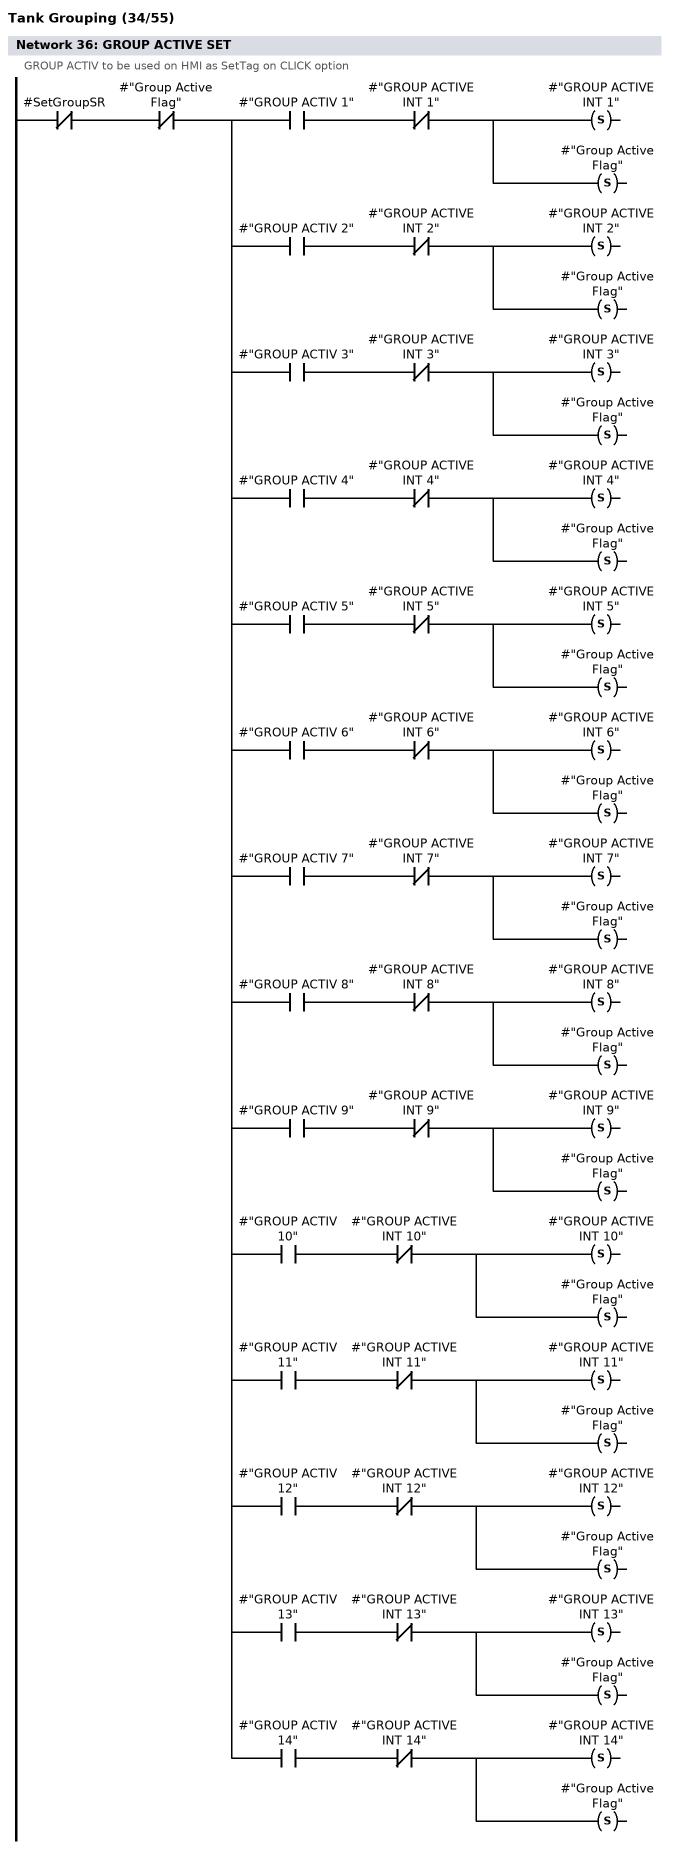
   RUNG wire#powerrail
      I_Contact( #SetGroupSR )
      I_Contact( #"Group Active Flag" )
      wire#w1
      Contact( #"GROUP ACTIV 1" )
      I_Contact( #"GROUP ACTIVE INT 1" )
      wire#w2
      S_Coil( #"GROUP ACTIVE INT 1" )
   END_RUNG
   RUNG wire#w2
      S_Coil( #"Group Active Flag" )
   END_RUNG
   RUNG wire#w1
      Contact( #"GROUP ACTIV 2" )
      I_Contact( #"GROUP ACTIVE INT 2" )
      wire#w3
      S_Coil( #"GROUP ACTIVE INT 2" )
   END_RUNG
   RUNG wire#w3
      S_Coil( #"Group Active Flag" )
   END_RUNG
   RUNG wire#w1
      Contact( #"GROUP ACTIV 3" )
      I_Contact( #"GROUP ACTIVE INT 3" )
      wire#w4
      S_Coil( #"GROUP ACTIVE INT 3" )
   END_RUNG
   RUNG wire#w4
      S_Coil( #"Group Active Flag" )
   END_RUNG
   RUNG wire#w1
      Contact( #"GROUP ACTIV 4" )
      I_Contact( #"GROUP ACTIVE INT 4" )
      wire#w5
      S_Coil( #"GROUP ACTIVE INT 4" )
   END_RUNG
   RUNG wire#w5
      S_Coil( #"Group Active Flag" )
   END_RUNG
   RUNG wire#w1
      Contact( #"GROUP ACTIV 5" )
      I_Contact( #"GROUP ACTIVE INT 5" )
      wire#w6
      S_Coil( #"GROUP ACTIVE INT 5" )
   END_RUNG
   RUNG wire#w6
      S_Coil( #"Group Active Flag" )
   END_RUNG
   RUNG wire#w1
      Contact( #"GROUP ACTIV 6" )
      I_Contact( #"GROUP ACTIVE INT 6" )
      wire#w7
      S_Coil( #"GROUP ACTIVE INT 6" )
   END_RUNG
   RUNG wire#w7
      S_Coil( #"Group Active Flag" )
   END_RUNG
   RUNG wire#w1
      Contact( #"GROUP ACTIV 7" )
      I_Contact( #"GROUP ACTIVE INT 7" )
      wire#w8
      S_Coil( #"GROUP ACTIVE INT 7" )
   END_RUNG
   RUNG wire#w8
      S_Coil( #"Group Active Flag" )
   END_RUNG
   RUNG wire#w1
      Contact( #"GROUP ACTIV 8" )
      I_Contact( #"GROUP ACTIVE INT 8" )
      wire#w9
      S_Coil( #"GROUP ACTIVE INT 8" )
   END_RUNG
   RUNG wire#w9
      S_Coil( #"Group Active Flag" )
   END_RUNG
   RUNG wire#w1
      Contact( #"GROUP ACTIV 9" )
      I_Contact( #"GROUP ACTIVE INT 9" )
      wire#w10
      S_Coil( #"GROUP ACTIVE INT 9" )
   END_RUNG
   RUNG wire#w10
      S_Coil( #"Group Active Flag" )
   END_RUNG
   RUNG wire#w1
      Contact( #"GROUP ACTIV 10" )
      I_Contact( #"GROUP ACTIVE INT 10" )
      wire#w11
      S_Coil( #"GROUP ACTIVE INT 10" )
   END_RUNG
   RUNG wire#w11
      S_Coil( #"Group Active Flag" )
   END_RUNG
   RUNG wire#w1
      Contact( #"GROUP ACTIV 11" )
      I_Contact( #"GROUP ACTIVE INT 11" )
      wire#w12
      S_Coil( #"GROUP ACTIVE INT 11" )
   END_RUNG
   RUNG wire#w12
      S_Coil( #"Group Active Flag" )
   END_RUNG
   RUNG wire#w1
      Contact( #"GROUP ACTIV 12" )
      I_Contact( #"GROUP ACTIVE INT 12" )
      wire#w13
      S_Coil( #"GROUP ACTIVE INT 12" )
   END_RUNG
   RUNG wire#w13
      S_Coil( #"Group Active Flag" )
   END_RUNG
   RUNG wire#w1
      Contact( #"GROUP ACTIV 13" )
      I_Contact( #"GROUP ACTIVE INT 13" )
      wire#w14
      S_Coil( #"GROUP ACTIVE INT 13" )
   END_RUNG
   RUNG wire#w14
      S_Coil( #"Group Active Flag" )
   END_RUNG
   RUNG wire#w1
      Contact( #"GROUP ACTIV 14" )
      I_Contact( #"GROUP ACTIVE INT 14" )
      wire#w15
      S_Coil( #"GROUP ACTIVE INT 14" )
   END_RUNG
   RUNG wire#w15
      S_Coil( #"Group Active Flag" )
   END_RUNG
   // the same network as SCL:
   #_w1 := NOT #SetGroupSR AND NOT #"Group Active Flag";
   #_w2 := #_w1 AND #"GROUP ACTIV 1" AND NOT #"GROUP ACTIVE INT 1";
   IF #_w2 THEN
       #"GROUP ACTIVE INT 1" := TRUE;
       #"Group Active Flag" := TRUE;
   END_IF;
   #_w3 := #_w1 AND #"GROUP ACTIV 2" AND NOT #"GROUP ACTIVE INT 2";
   IF #_w3 THEN
       #"GROUP ACTIVE INT 2" := TRUE;
       #"Group Active Flag" := TRUE;
   END_IF;
   #_w4 := #_w1 AND #"GROUP ACTIV 3" AND NOT #"GROUP ACTIVE INT 3";
   IF #_w4 THEN
       #"GROUP ACTIVE INT 3" := TRUE;
       #"Group Active Flag" := TRUE;
   END_IF;
   #_w5 := #_w1 AND #"GROUP ACTIV 4" AND NOT #"GROUP ACTIVE INT 4";
   IF #_w5 THEN
       #"GROUP ACTIVE INT 4" := TRUE;
       #"Group Active Flag" := TRUE;
   END_IF;
   #_w6 := #_w1 AND #"GROUP ACTIV 5" AND NOT #"GROUP ACTIVE INT 5";
   IF #_w6 THEN
       #"GROUP ACTIVE INT 5" := TRUE;
       #"Group Active Flag" := TRUE;
   END_IF;
   #_w7 := #_w1 AND #"GROUP ACTIV 6" AND NOT #"GROUP ACTIVE INT 6";
   IF #_w7 THEN
       #"GROUP ACTIVE INT 6" := TRUE;
       #"Group Active Flag" := TRUE;
   END_IF;
   #_w8 := #_w1 AND #"GROUP ACTIV 7" AND NOT #"GROUP ACTIVE INT 7";
   IF #_w8 THEN
       #"GROUP ACTIVE INT 7" := TRUE;
       #"Group Active Flag" := TRUE;
   END_IF;
   #_w9 := #_w1 AND #"GROUP ACTIV 8" AND NOT #"GROUP ACTIVE INT 8";
   IF #_w9 THEN
       #"GROUP ACTIVE INT 8" := TRUE;
       #"Group Active Flag" := TRUE;
   END_IF;
   #_w10 := #_w1 AND #"GROUP ACTIV 9" AND NOT #"GROUP ACTIVE INT 9";
   IF #_w10 THEN
       #"GROUP ACTIVE INT 9" := TRUE;
       #"Group Active Flag" := TRUE;
   END_IF;
   #_w11 := #_w1 AND #"GROUP ACTIV 10" AND NOT #"GROUP ACTIVE INT 10";
   IF #_w11 THEN
       #"GROUP ACTIVE INT 10" := TRUE;
       #"Group Active Flag" := TRUE;
   END_IF;
   #_w12 := #_w1 AND #"GROUP ACTIV 11" AND NOT #"GROUP ACTIVE INT 11";
   IF #_w12 THEN
       #"GROUP ACTIVE INT 11" := TRUE;
       #"Group Active Flag" := TRUE;
   END_IF;
   #_w13 := #_w1 AND #"GROUP ACTIV 12" AND NOT #"GROUP ACTIVE INT 12";
   IF #_w13 THEN
       #"GROUP ACTIVE INT 12" := TRUE;
       #"Group Active Flag" := TRUE;
   END_IF;
   #_w14 := #_w1 AND #"GROUP ACTIV 13" AND NOT #"GROUP ACTIVE INT 13";
   IF #_w14 THEN
       #"GROUP ACTIVE INT 13" := TRUE;
       #"Group Active Flag" := TRUE;
   END_IF;
   #_w15 := #_w1 AND #"GROUP ACTIV 14" AND NOT #"GROUP ACTIVE INT 14";
   IF #_w15 THEN
       #"GROUP ACTIVE INT 14" := TRUE;
       #"Group Active Flag" := TRUE;
   END_IF;
END_REGION

REGION Network 37: Group Active Flag Reset
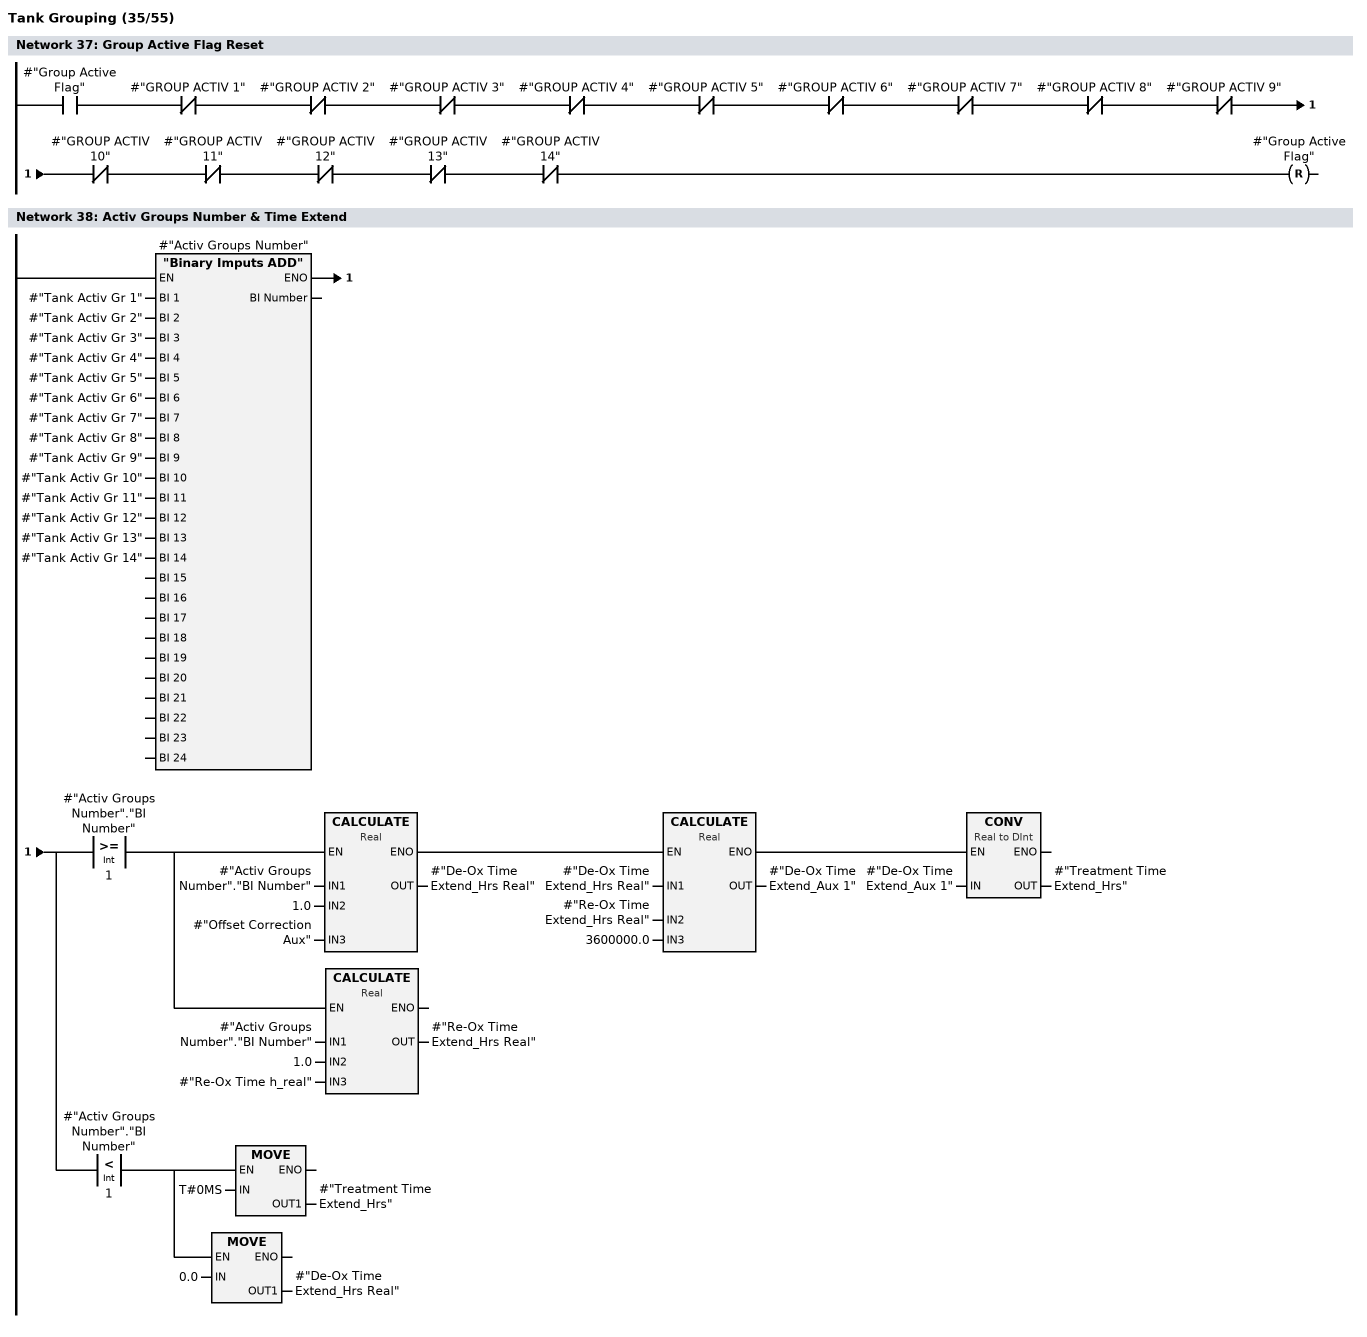
   RUNG wire#powerrail
      Contact( #"Group Active Flag" )
      I_Contact( #"GROUP ACTIV 1" )
      I_Contact( #"GROUP ACTIV 2" )
      I_Contact( #"GROUP ACTIV 3" )
      I_Contact( #"GROUP ACTIV 4" )
      I_Contact( #"GROUP ACTIV 5" )
      I_Contact( #"GROUP ACTIV 6" )
      I_Contact( #"GROUP ACTIV 7" )
      I_Contact( #"GROUP ACTIV 8" )
      I_Contact( #"GROUP ACTIV 9" )
      I_Contact( #"GROUP ACTIV 10" )
      I_Contact( #"GROUP ACTIV 11" )
      I_Contact( #"GROUP ACTIV 12" )
      I_Contact( #"GROUP ACTIV 13" )
      I_Contact( #"GROUP ACTIV 14" )
      R_Coil( #"Group Active Flag" )
   END_RUNG
   // the same network as SCL:
   IF #"Group Active Flag" AND NOT #"GROUP ACTIV 1" AND NOT #"GROUP ACTIV 2" AND NOT #"GROUP ACTIV 3" AND NOT #"GROUP ACTIV 4" AND NOT #"GROUP ACTIV 5" AND NOT #"GROUP ACTIV 6" AND NOT #"GROUP ACTIV 7" AND NOT #"GROUP ACTIV 8" AND NOT #"GROUP ACTIV 9" AND NOT #"GROUP ACTIV 10" AND NOT #"GROUP ACTIV 11" AND NOT #"GROUP ACTIV 12" AND NOT #"GROUP ACTIV 13" AND NOT #"GROUP ACTIV 14" THEN
       #"Group Active Flag" := FALSE;
   END_IF;
END_REGION

REGION Network 38: Activ Groups Number & Time Extend
   RUNG wire#powerrail
      #"Activ Groups Number"("BI 1" := #"Tank Activ Gr 1", "BI 2" := #"Tank Activ Gr 2", "BI 3" := #"Tank Activ Gr 3", "BI 4" := #"Tank Activ Gr 4", "BI 5" := #"Tank Activ Gr 5", "BI 6" := #"Tank Activ Gr 6", "BI 7" := #"Tank Activ Gr 7", "BI 8" := #"Tank Activ Gr 8", "BI 9" := #"Tank Activ Gr 9", "BI 10" := #"Tank Activ Gr 10", "BI 11" := #"Tank Activ Gr 11", "BI 12" := #"Tank Activ Gr 12", "BI 13" := #"Tank Activ Gr 13", "BI 14" := #"Tank Activ Gr 14", "BI 15" :=, "BI 16" :=, "BI 17" :=, "BI 18" :=, "BI 19" :=, "BI 20" :=, "BI 21" :=, "BI 22" :=, "BI 23" :=, "BI 24" :=, "BI Number" =>)
      wire#w1
      { S7_Templates := "SrcType := Int" } GE_Contact(in1 := #"Activ Groups Number"."BI Number", in2 := 1)
      wire#w2
      { S7_Templates := "SrcType := Real"; S7_Expression := "IN3*(IN1-IN2)" } Calculate(in1 := #"Activ Groups Number"."BI Number", in2 := 1.0, in3 := #"Offset Correction Aux", out => #"De-Ox Time Extend_Hrs Real")
      { S7_Templates := "SrcType := Real"; S7_Expression := "(IN1+IN2)*IN3" } Calculate(in1 := #"De-Ox Time Extend_Hrs Real", in2 := #"Re-Ox Time Extend_Hrs Real", in3 := 3600000.0, out => #"De-Ox Time Extend_Aux 1")
      { S7_Templates := "[SrcType := Real, DestType := DInt]" } Convert(in := #"De-Ox Time Extend_Aux 1", out => #"Treatment Time Extend_Hrs")
   END_RUNG
   RUNG wire#w2
      { S7_Templates := "SrcType := Real"; S7_Expression := "IN3*(IN1-IN2)" } Calculate(in1 := #"Activ Groups Number"."BI Number", in2 := 1.0, in3 := #"Re-Ox Time h_real", out => #"Re-Ox Time Extend_Hrs Real")
   END_RUNG
   RUNG wire#w1
      { S7_Templates := "SrcType := Int" } LT_Contact(in1 := #"Activ Groups Number"."BI Number", in2 := 1)
      wire#w3
      Move(in := T#0MS, out1 => #"Treatment Time Extend_Hrs")
   END_RUNG
   RUNG wire#w3
      Move(in := 0.0, out1 => #"De-Ox Time Extend_Hrs Real")
   END_RUNG
   // the same network as SCL:
   #"Activ Groups Number"("BI 1" := #"Tank Activ Gr 1",   // "Binary Imputs ADD"
                          "BI 2" := #"Tank Activ Gr 2",
                          "BI 3" := #"Tank Activ Gr 3",
                          "BI 4" := #"Tank Activ Gr 4",
                          "BI 5" := #"Tank Activ Gr 5",
                          "BI 6" := #"Tank Activ Gr 6",
                          "BI 7" := #"Tank Activ Gr 7",
                          "BI 8" := #"Tank Activ Gr 8",
                          "BI 9" := #"Tank Activ Gr 9",
                          "BI 10" := #"Tank Activ Gr 10",
                          "BI 11" := #"Tank Activ Gr 11",
                          "BI 12" := #"Tank Activ Gr 12",
                          "BI 13" := #"Tank Activ Gr 13",
                          "BI 14" := #"Tank Activ Gr 14",
                          ENO => #_w1);
   IF #_w1 AND (#"Activ Groups Number"."BI Number" >= 1) THEN
       #"De-Ox Time Extend_Hrs Real" := #"Offset Correction Aux"*(#"Activ Groups Number"."BI Number"-1.0);
       #"De-Ox Time Extend_Aux 1" := (#"De-Ox Time Extend_Hrs Real"+#"Re-Ox Time Extend_Hrs Real")*3600000.0;
       #"Treatment Time Extend_Hrs" := REAL_TO_DINT(#"De-Ox Time Extend_Aux 1");
       #"Re-Ox Time Extend_Hrs Real" := #"Re-Ox Time h_real"*(#"Activ Groups Number"."BI Number"-1.0);
   END_IF;
   IF #_w1 AND (#"Activ Groups Number"."BI Number" < 1) THEN
       #"Treatment Time Extend_Hrs" := T#0MS;
       #"De-Ox Time Extend_Hrs Real" := 0.0;
   END_IF;
END_REGION

REGION Network 39: GROUP ACTIVE RESET
   // GROUP ACTIV to be used on HMI as SetTag on CLICK option
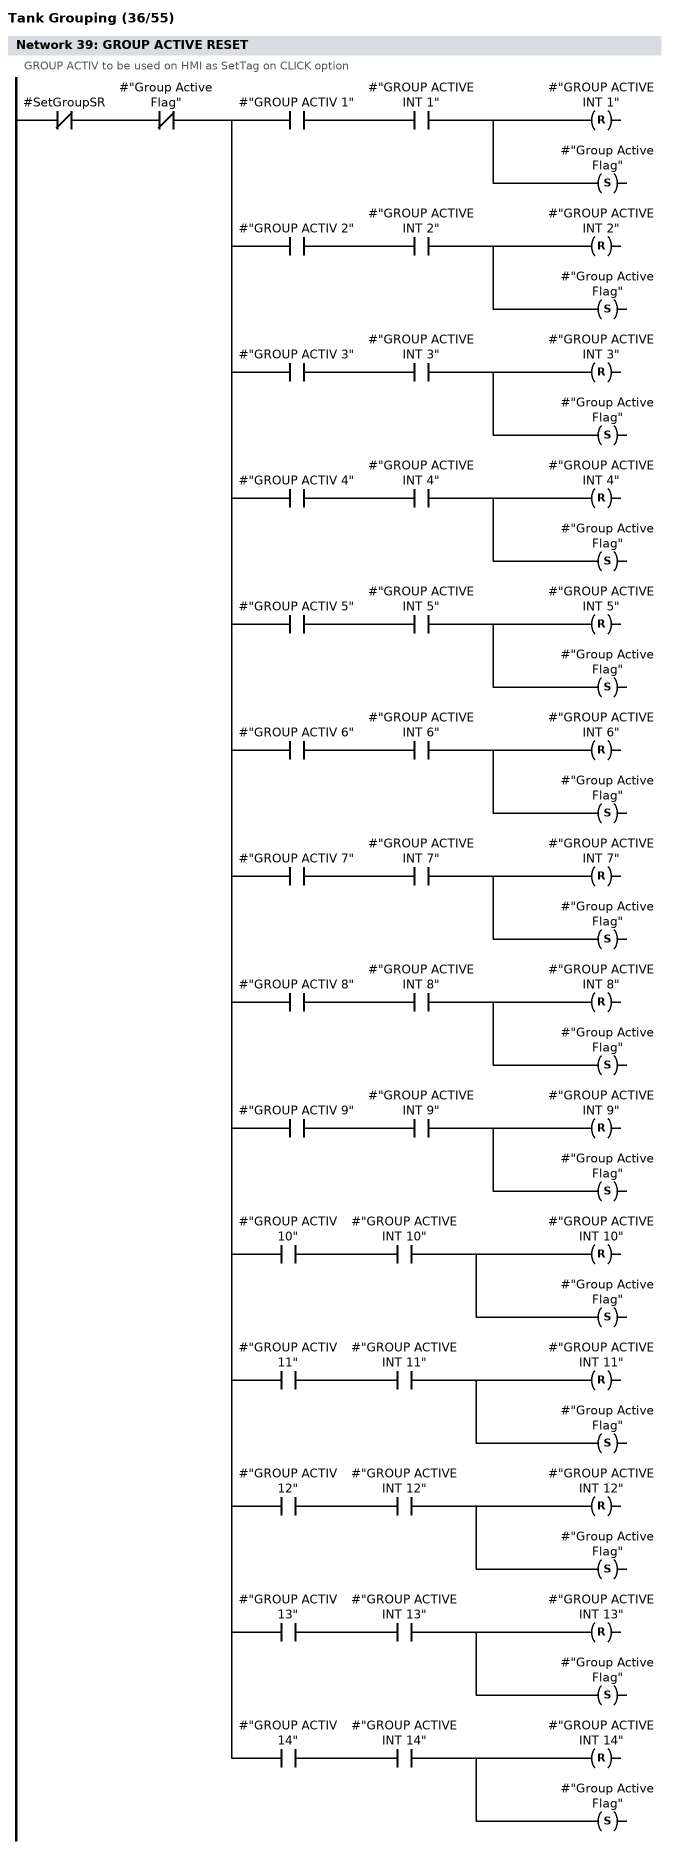
   RUNG wire#powerrail
      I_Contact( #SetGroupSR )
      I_Contact( #"Group Active Flag" )
      wire#w1
      Contact( #"GROUP ACTIV 1" )
      Contact( #"GROUP ACTIVE INT 1" )
      wire#w2
      R_Coil( #"GROUP ACTIVE INT 1" )
   END_RUNG
   RUNG wire#w2
      S_Coil( #"Group Active Flag" )
   END_RUNG
   RUNG wire#w1
      Contact( #"GROUP ACTIV 2" )
      Contact( #"GROUP ACTIVE INT 2" )
      wire#w3
      R_Coil( #"GROUP ACTIVE INT 2" )
   END_RUNG
   RUNG wire#w3
      S_Coil( #"Group Active Flag" )
   END_RUNG
   RUNG wire#w1
      Contact( #"GROUP ACTIV 3" )
      Contact( #"GROUP ACTIVE INT 3" )
      wire#w4
      R_Coil( #"GROUP ACTIVE INT 3" )
   END_RUNG
   RUNG wire#w4
      S_Coil( #"Group Active Flag" )
   END_RUNG
   RUNG wire#w1
      Contact( #"GROUP ACTIV 4" )
      Contact( #"GROUP ACTIVE INT 4" )
      wire#w5
      R_Coil( #"GROUP ACTIVE INT 4" )
   END_RUNG
   RUNG wire#w5
      S_Coil( #"Group Active Flag" )
   END_RUNG
   RUNG wire#w1
      Contact( #"GROUP ACTIV 5" )
      Contact( #"GROUP ACTIVE INT 5" )
      wire#w6
      R_Coil( #"GROUP ACTIVE INT 5" )
   END_RUNG
   RUNG wire#w6
      S_Coil( #"Group Active Flag" )
   END_RUNG
   RUNG wire#w1
      Contact( #"GROUP ACTIV 6" )
      Contact( #"GROUP ACTIVE INT 6" )
      wire#w7
      R_Coil( #"GROUP ACTIVE INT 6" )
   END_RUNG
   RUNG wire#w7
      S_Coil( #"Group Active Flag" )
   END_RUNG
   RUNG wire#w1
      Contact( #"GROUP ACTIV 7" )
      Contact( #"GROUP ACTIVE INT 7" )
      wire#w8
      R_Coil( #"GROUP ACTIVE INT 7" )
   END_RUNG
   RUNG wire#w8
      S_Coil( #"Group Active Flag" )
   END_RUNG
   RUNG wire#w1
      Contact( #"GROUP ACTIV 8" )
      Contact( #"GROUP ACTIVE INT 8" )
      wire#w9
      R_Coil( #"GROUP ACTIVE INT 8" )
   END_RUNG
   RUNG wire#w9
      S_Coil( #"Group Active Flag" )
   END_RUNG
   RUNG wire#w1
      Contact( #"GROUP ACTIV 9" )
      Contact( #"GROUP ACTIVE INT 9" )
      wire#w10
      R_Coil( #"GROUP ACTIVE INT 9" )
   END_RUNG
   RUNG wire#w10
      S_Coil( #"Group Active Flag" )
   END_RUNG
   RUNG wire#w1
      Contact( #"GROUP ACTIV 10" )
      Contact( #"GROUP ACTIVE INT 10" )
      wire#w11
      R_Coil( #"GROUP ACTIVE INT 10" )
   END_RUNG
   RUNG wire#w11
      S_Coil( #"Group Active Flag" )
   END_RUNG
   RUNG wire#w1
      Contact( #"GROUP ACTIV 11" )
      Contact( #"GROUP ACTIVE INT 11" )
      wire#w12
      R_Coil( #"GROUP ACTIVE INT 11" )
   END_RUNG
   RUNG wire#w12
      S_Coil( #"Group Active Flag" )
   END_RUNG
   RUNG wire#w1
      Contact( #"GROUP ACTIV 12" )
      Contact( #"GROUP ACTIVE INT 12" )
      wire#w13
      R_Coil( #"GROUP ACTIVE INT 12" )
   END_RUNG
   RUNG wire#w13
      S_Coil( #"Group Active Flag" )
   END_RUNG
   RUNG wire#w1
      Contact( #"GROUP ACTIV 13" )
      Contact( #"GROUP ACTIVE INT 13" )
      wire#w14
      R_Coil( #"GROUP ACTIVE INT 13" )
   END_RUNG
   RUNG wire#w14
      S_Coil( #"Group Active Flag" )
   END_RUNG
   RUNG wire#w1
      Contact( #"GROUP ACTIV 14" )
      Contact( #"GROUP ACTIVE INT 14" )
      wire#w15
      R_Coil( #"GROUP ACTIVE INT 14" )
   END_RUNG
   RUNG wire#w15
      S_Coil( #"Group Active Flag" )
   END_RUNG
   // the same network as SCL:
   #_w1 := NOT #SetGroupSR AND NOT #"Group Active Flag";
   #_w2 := #_w1 AND #"GROUP ACTIV 1" AND #"GROUP ACTIVE INT 1";
   IF #_w2 THEN
       #"GROUP ACTIVE INT 1" := FALSE;
       #"Group Active Flag" := TRUE;
   END_IF;
   #_w3 := #_w1 AND #"GROUP ACTIV 2" AND #"GROUP ACTIVE INT 2";
   IF #_w3 THEN
       #"GROUP ACTIVE INT 2" := FALSE;
       #"Group Active Flag" := TRUE;
   END_IF;
   #_w4 := #_w1 AND #"GROUP ACTIV 3" AND #"GROUP ACTIVE INT 3";
   IF #_w4 THEN
       #"GROUP ACTIVE INT 3" := FALSE;
       #"Group Active Flag" := TRUE;
   END_IF;
   #_w5 := #_w1 AND #"GROUP ACTIV 4" AND #"GROUP ACTIVE INT 4";
   IF #_w5 THEN
       #"GROUP ACTIVE INT 4" := FALSE;
       #"Group Active Flag" := TRUE;
   END_IF;
   #_w6 := #_w1 AND #"GROUP ACTIV 5" AND #"GROUP ACTIVE INT 5";
   IF #_w6 THEN
       #"GROUP ACTIVE INT 5" := FALSE;
       #"Group Active Flag" := TRUE;
   END_IF;
   #_w7 := #_w1 AND #"GROUP ACTIV 6" AND #"GROUP ACTIVE INT 6";
   IF #_w7 THEN
       #"GROUP ACTIVE INT 6" := FALSE;
       #"Group Active Flag" := TRUE;
   END_IF;
   #_w8 := #_w1 AND #"GROUP ACTIV 7" AND #"GROUP ACTIVE INT 7";
   IF #_w8 THEN
       #"GROUP ACTIVE INT 7" := FALSE;
       #"Group Active Flag" := TRUE;
   END_IF;
   #_w9 := #_w1 AND #"GROUP ACTIV 8" AND #"GROUP ACTIVE INT 8";
   IF #_w9 THEN
       #"GROUP ACTIVE INT 8" := FALSE;
       #"Group Active Flag" := TRUE;
   END_IF;
   #_w10 := #_w1 AND #"GROUP ACTIV 9" AND #"GROUP ACTIVE INT 9";
   IF #_w10 THEN
       #"GROUP ACTIVE INT 9" := FALSE;
       #"Group Active Flag" := TRUE;
   END_IF;
   #_w11 := #_w1 AND #"GROUP ACTIV 10" AND #"GROUP ACTIVE INT 10";
   IF #_w11 THEN
       #"GROUP ACTIVE INT 10" := FALSE;
       #"Group Active Flag" := TRUE;
   END_IF;
   #_w12 := #_w1 AND #"GROUP ACTIV 11" AND #"GROUP ACTIVE INT 11";
   IF #_w12 THEN
       #"GROUP ACTIVE INT 11" := FALSE;
       #"Group Active Flag" := TRUE;
   END_IF;
   #_w13 := #_w1 AND #"GROUP ACTIV 12" AND #"GROUP ACTIVE INT 12";
   IF #_w13 THEN
       #"GROUP ACTIVE INT 12" := FALSE;
       #"Group Active Flag" := TRUE;
   END_IF;
   #_w14 := #_w1 AND #"GROUP ACTIV 13" AND #"GROUP ACTIVE INT 13";
   IF #_w14 THEN
       #"GROUP ACTIVE INT 13" := FALSE;
       #"Group Active Flag" := TRUE;
   END_IF;
   #_w15 := #_w1 AND #"GROUP ACTIV 14" AND #"GROUP ACTIVE INT 14";
   IF #_w15 THEN
       #"GROUP ACTIVE INT 14" := FALSE;
       #"Group Active Flag" := TRUE;
   END_IF;
END_REGION

REGION Network 40: Tank Treatment Offset
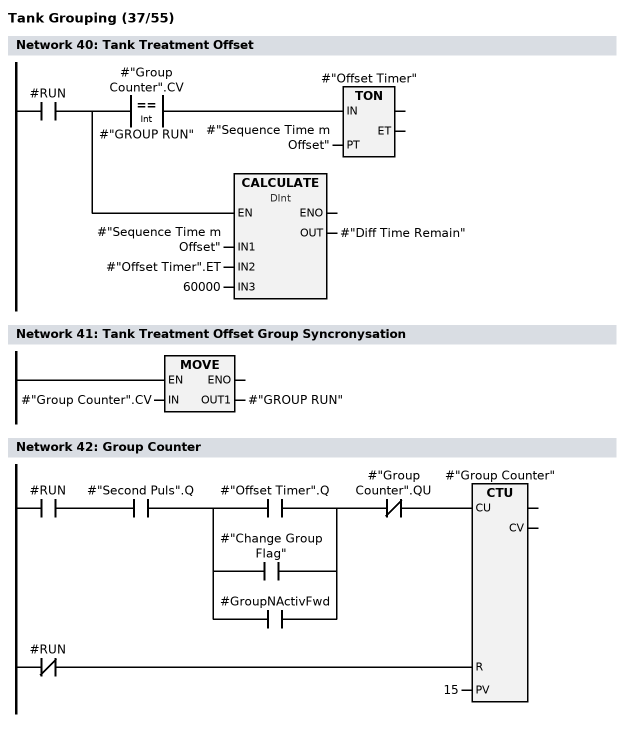
   #"Offset Timer"(IN := #RUN AND (#"Group Counter".CV = #"GROUP RUN"), PT := #"Sequence Time m Offset");   // TON
   IF #RUN THEN #"Diff Time Remain" := (#"Sequence Time m Offset"-#"Offset Timer".ET)/60000; END_IF;
END_REGION

REGION Network 41: Tank Treatment Offset Group Syncronysation
   RUNG wire#powerrail
      Move(in := #"Group Counter".CV, out1 => #"GROUP RUN")
   END_RUNG
   // the same network as SCL:
   #"GROUP RUN" := #"Group Counter".CV;
END_REGION

REGION Network 42: Group Counter
   #"Group Counter"(CU := #RUN AND #"Second Puls".Q AND (#"Offset Timer".Q OR #"Change Group Flag" OR #GroupNActivFwd) AND NOT #"Group Counter".QU,   // CTU
                    R := NOT #RUN,
                    PV := 15);
END_REGION

REGION Network 43: RUN GROUP
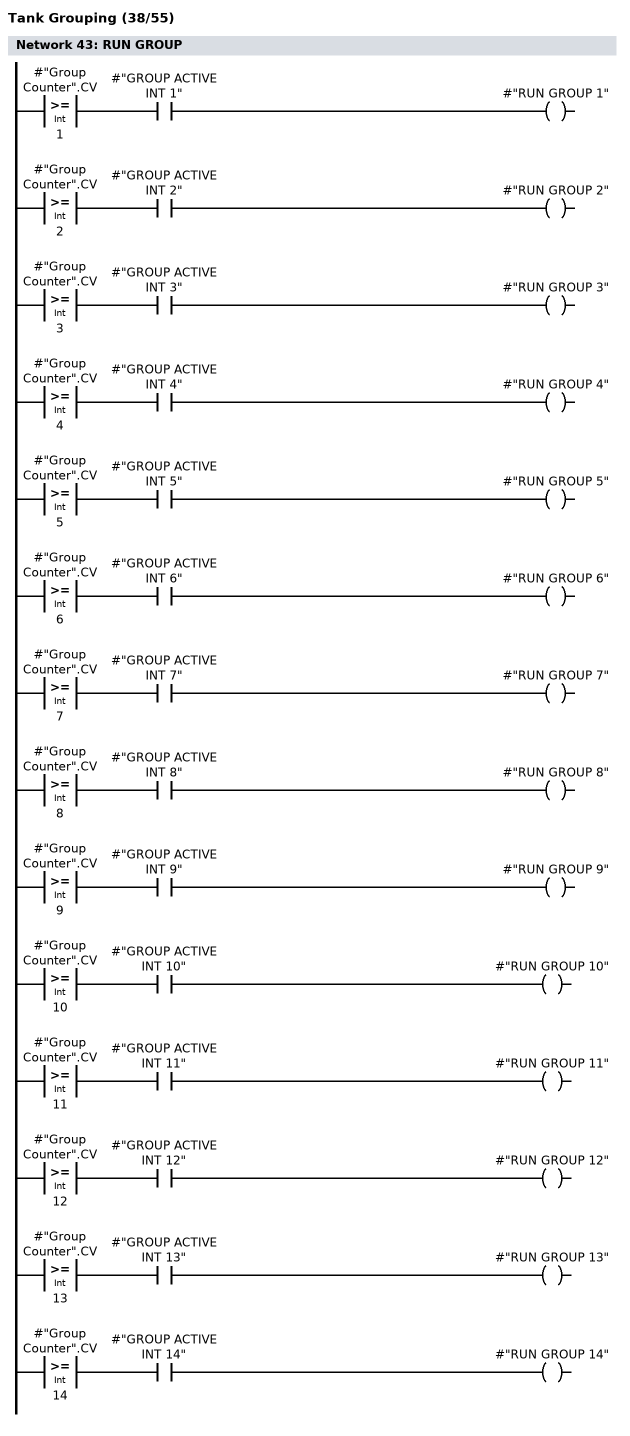
   RUNG wire#powerrail
      { S7_Templates := "SrcType := Int" } GE_Contact(in1 := #"Group Counter".CV, in2 := 1)
      Contact( #"GROUP ACTIVE INT 1" )
      Coil( #"RUN GROUP 1" )
   END_RUNG
   RUNG wire#powerrail
      { S7_Templates := "SrcType := Int" } GE_Contact(in1 := #"Group Counter".CV, in2 := 2)
      Contact( #"GROUP ACTIVE INT 2" )
      Coil( #"RUN GROUP 2" )
   END_RUNG
   RUNG wire#powerrail
      { S7_Templates := "SrcType := Int" } GE_Contact(in1 := #"Group Counter".CV, in2 := 3)
      Contact( #"GROUP ACTIVE INT 3" )
      Coil( #"RUN GROUP 3" )
   END_RUNG
   RUNG wire#powerrail
      { S7_Templates := "SrcType := Int" } GE_Contact(in1 := #"Group Counter".CV, in2 := 4)
      Contact( #"GROUP ACTIVE INT 4" )
      Coil( #"RUN GROUP 4" )
   END_RUNG
   RUNG wire#powerrail
      { S7_Templates := "SrcType := Int" } GE_Contact(in1 := #"Group Counter".CV, in2 := 5)
      Contact( #"GROUP ACTIVE INT 5" )
      Coil( #"RUN GROUP 5" )
   END_RUNG
   RUNG wire#powerrail
      { S7_Templates := "SrcType := Int" } GE_Contact(in1 := #"Group Counter".CV, in2 := 6)
      Contact( #"GROUP ACTIVE INT 6" )
      Coil( #"RUN GROUP 6" )
   END_RUNG
   RUNG wire#powerrail
      { S7_Templates := "SrcType := Int" } GE_Contact(in1 := #"Group Counter".CV, in2 := 7)
      Contact( #"GROUP ACTIVE INT 7" )
      Coil( #"RUN GROUP 7" )
   END_RUNG
   RUNG wire#powerrail
      { S7_Templates := "SrcType := Int" } GE_Contact(in1 := #"Group Counter".CV, in2 := 8)
      Contact( #"GROUP ACTIVE INT 8" )
      Coil( #"RUN GROUP 8" )
   END_RUNG
   RUNG wire#powerrail
      { S7_Templates := "SrcType := Int" } GE_Contact(in1 := #"Group Counter".CV, in2 := 9)
      Contact( #"GROUP ACTIVE INT 9" )
      Coil( #"RUN GROUP 9" )
   END_RUNG
   RUNG wire#powerrail
      { S7_Templates := "SrcType := Int" } GE_Contact(in1 := #"Group Counter".CV, in2 := 10)
      Contact( #"GROUP ACTIVE INT 10" )
      Coil( #"RUN GROUP 10" )
   END_RUNG
   RUNG wire#powerrail
      { S7_Templates := "SrcType := Int" } GE_Contact(in1 := #"Group Counter".CV, in2 := 11)
      Contact( #"GROUP ACTIVE INT 11" )
      Coil( #"RUN GROUP 11" )
   END_RUNG
   RUNG wire#powerrail
      { S7_Templates := "SrcType := Int" } GE_Contact(in1 := #"Group Counter".CV, in2 := 12)
      Contact( #"GROUP ACTIVE INT 12" )
      Coil( #"RUN GROUP 12" )
   END_RUNG
   RUNG wire#powerrail
      { S7_Templates := "SrcType := Int" } GE_Contact(in1 := #"Group Counter".CV, in2 := 13)
      Contact( #"GROUP ACTIVE INT 13" )
      Coil( #"RUN GROUP 13" )
   END_RUNG
   RUNG wire#powerrail
      { S7_Templates := "SrcType := Int" } GE_Contact(in1 := #"Group Counter".CV, in2 := 14)
      Contact( #"GROUP ACTIVE INT 14" )
      Coil( #"RUN GROUP 14" )
   END_RUNG
   // the same network as SCL:
   #"RUN GROUP 1" := (#"Group Counter".CV >= 1) AND #"GROUP ACTIVE INT 1";
   #"RUN GROUP 2" := (#"Group Counter".CV >= 2) AND #"GROUP ACTIVE INT 2";
   #"RUN GROUP 3" := (#"Group Counter".CV >= 3) AND #"GROUP ACTIVE INT 3";
   #"RUN GROUP 4" := (#"Group Counter".CV >= 4) AND #"GROUP ACTIVE INT 4";
   #"RUN GROUP 5" := (#"Group Counter".CV >= 5) AND #"GROUP ACTIVE INT 5";
   #"RUN GROUP 6" := (#"Group Counter".CV >= 6) AND #"GROUP ACTIVE INT 6";
   #"RUN GROUP 7" := (#"Group Counter".CV >= 7) AND #"GROUP ACTIVE INT 7";
   #"RUN GROUP 8" := (#"Group Counter".CV >= 8) AND #"GROUP ACTIVE INT 8";
   #"RUN GROUP 9" := (#"Group Counter".CV >= 9) AND #"GROUP ACTIVE INT 9";
   #"RUN GROUP 10" := (#"Group Counter".CV >= 10) AND #"GROUP ACTIVE INT 10";
   #"RUN GROUP 11" := (#"Group Counter".CV >= 11) AND #"GROUP ACTIVE INT 11";
   #"RUN GROUP 12" := (#"Group Counter".CV >= 12) AND #"GROUP ACTIVE INT 12";
   #"RUN GROUP 13" := (#"Group Counter".CV >= 13) AND #"GROUP ACTIVE INT 13";
   #"RUN GROUP 14" := (#"Group Counter".CV >= 14) AND #"GROUP ACTIVE INT 14";
END_REGION

REGION Network 44: RUN GROUP INACTIV MOVE FORWARD
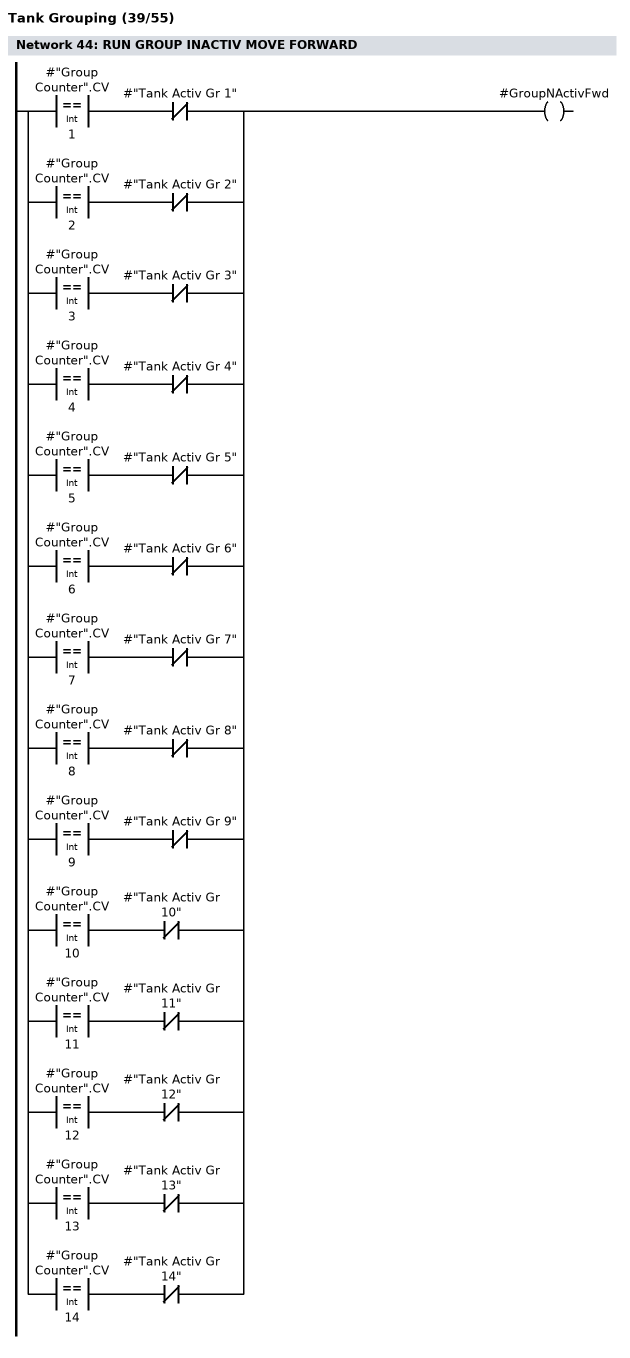
   RUNG wire#powerrail
      { S7_Templates := "SrcType := Int" } EQ_Contact(in1 := #"Group Counter".CV, in2 := 1)
      I_Contact( #"Tank Activ Gr 1" )
      wire#w1
      Coil( #GroupNActivFwd )
   END_RUNG
   RUNG wire#powerrail
      { S7_Templates := "SrcType := Int" } EQ_Contact(in1 := #"Group Counter".CV, in2 := 2)
      I_Contact( #"Tank Activ Gr 2" )
   END_RUNG wire#w1
   RUNG wire#powerrail
      { S7_Templates := "SrcType := Int" } EQ_Contact(in1 := #"Group Counter".CV, in2 := 3)
      I_Contact( #"Tank Activ Gr 3" )
   END_RUNG wire#w1
   RUNG wire#powerrail
      { S7_Templates := "SrcType := Int" } EQ_Contact(in1 := #"Group Counter".CV, in2 := 4)
      I_Contact( #"Tank Activ Gr 4" )
   END_RUNG wire#w1
   RUNG wire#powerrail
      { S7_Templates := "SrcType := Int" } EQ_Contact(in1 := #"Group Counter".CV, in2 := 5)
      I_Contact( #"Tank Activ Gr 5" )
   END_RUNG wire#w1
   RUNG wire#powerrail
      { S7_Templates := "SrcType := Int" } EQ_Contact(in1 := #"Group Counter".CV, in2 := 6)
      I_Contact( #"Tank Activ Gr 6" )
   END_RUNG wire#w1
   RUNG wire#powerrail
      { S7_Templates := "SrcType := Int" } EQ_Contact(in1 := #"Group Counter".CV, in2 := 7)
      I_Contact( #"Tank Activ Gr 7" )
   END_RUNG wire#w1
   RUNG wire#powerrail
      { S7_Templates := "SrcType := Int" } EQ_Contact(in1 := #"Group Counter".CV, in2 := 8)
      I_Contact( #"Tank Activ Gr 8" )
   END_RUNG wire#w1
   RUNG wire#powerrail
      { S7_Templates := "SrcType := Int" } EQ_Contact(in1 := #"Group Counter".CV, in2 := 9)
      I_Contact( #"Tank Activ Gr 9" )
   END_RUNG wire#w1
   RUNG wire#powerrail
      { S7_Templates := "SrcType := Int" } EQ_Contact(in1 := #"Group Counter".CV, in2 := 10)
      I_Contact( #"Tank Activ Gr 10" )
   END_RUNG wire#w1
   RUNG wire#powerrail
      { S7_Templates := "SrcType := Int" } EQ_Contact(in1 := #"Group Counter".CV, in2 := 11)
      I_Contact( #"Tank Activ Gr 11" )
   END_RUNG wire#w1
   RUNG wire#powerrail
      { S7_Templates := "SrcType := Int" } EQ_Contact(in1 := #"Group Counter".CV, in2 := 12)
      I_Contact( #"Tank Activ Gr 12" )
   END_RUNG wire#w1
   RUNG wire#powerrail
      { S7_Templates := "SrcType := Int" } EQ_Contact(in1 := #"Group Counter".CV, in2 := 13)
      I_Contact( #"Tank Activ Gr 13" )
   END_RUNG wire#w1
   RUNG wire#powerrail
      { S7_Templates := "SrcType := Int" } EQ_Contact(in1 := #"Group Counter".CV, in2 := 14)
      I_Contact( #"Tank Activ Gr 14" )
   END_RUNG wire#w1
   // the same network as SCL:
   #GroupNActivFwd := ((#"Group Counter".CV = 1) AND NOT #"Tank Activ Gr 1") OR ((#"Group Counter".CV = 2) AND NOT #"Tank Activ Gr 2") OR ((#"Group Counter".CV = 3) AND NOT #"Tank Activ Gr 3") OR ((#"Group Counter".CV = 4) AND NOT #"Tank Activ Gr 4") OR ((#"Group Counter".CV = 5) AND NOT #"Tank Activ Gr 5") OR ((#"Group Counter".CV = 6) AND NOT #"Tank Activ Gr 6") OR ((#"Group Counter".CV = 7) AND NOT #"Tank Activ Gr 7") OR ((#"Group Counter".CV = 8) AND NOT #"Tank Activ Gr 8") OR ((#"Group Counter".CV = 9) AND NOT #"Tank Activ Gr 9") OR ((#"Group Counter".CV = 10) AND NOT #"Tank Activ Gr 10") OR ((#"Group Counter".CV = 11) AND NOT #"Tank Activ Gr 11") OR ((#"Group Counter".CV = 12) AND NOT #"Tank Activ Gr 12") OR ((#"Group Counter".CV = 13) AND NOT #"Tank Activ Gr 13") OR ((#"Group Counter".CV = 14) AND NOT #"Tank Activ Gr 14");
END_REGION

REGION Network 45: Change Group Flag